
   IF #statErrorUserCleared = TRUE 
   THEN

       REGION Program

           //copy new value
           #statValues[0] := #statValues[1]; // -> n-2
           #statValues[1] := #statValues[2]; // -> n-1
           #statValues[2] := #statValues[3]; // -> n
           #statValues[3] := #statValues[4]; // -> n+1
           #statValues[4] := #value;         // -> n+2

           IF #statCount < 4
           THEN
               #status:= #STATUS_NOT_ENOUGH_VALUES;
               #statCount += 1;
               #statErrorAutoCleared := true;
           ELSE
               //calculate new smoothed value 
               //ẏ(n)=1/12deltaT*(y(n-2)-8y(n-1)+8y(n+1)-y(n+2))
               //1/12deltaT = 
               #statDerivatedValue := LREAL_TO_REAL(1.0 / (12.0*#deltaT)) * (#statValues[0] -8 * #statValues[1] + 8 * #statValues[3] - #statValues[4]);
               #statDone := true;
           END_IF;

       END_REGION
   END_IF;

   //----------------------------------------------------------------------------------------------
   //Write ouputs and error handling
   //----------------------------------------------------------------------------------------------
   //Error occured in request
   IF #statErrorAutoCleared
   THEN
       #statDone := FALSE;
       #statErrorUserCleared := FALSE;
       //Request finished
   ELSIF #statDone
   THEN
       #statErrorUserCleared := FALSE;
       #statErrorAutoCleared := FALSE;
       #status := #STATUS_EXECUTION_FINISHED;
       #derivatedValue := #statDerivatedValue;
       //Request in execution
   ELSE
       #status := #STATUS_SUBSEQUENT_CALL;
   END_IF;

   //Write static values to outputs
   #valid := #statDone;
   #busy := #statErrorUserCleared;
   #error := #statErrorAutoCleared;
   //----------------------------------------------------------------------------------------------

   //=============================================================================

   //----------------------------------------------------------------------------------------------
   //Check if FB is disabled
   IF NOT #enable
     AND #statEnableOld
   THEN

     //Error outputs are reset with falling edge of enable input
     #statErrorUserCleared := FALSE;
     #statErrorAutoCleared := FALSE;
     #error := FALSE;
     #status := #STATUS_NO_CALL;

     //Enable and busy are reset with falling edge of enable input
     #busy := FALSE;
     #busy := FALSE;

     //Set old value of enable for edge detection and end execution
     #statEnableOld := #enable;
     RETURN;

     //Check if FB is enabled
   ELSIF #enable
     AND NOT #statEnableOld
   THEN
     //reset static values
     #statCount := 0;
     #statValues[0] := 0.0;
     #statValues[1] := 0.0;
     #statValues[2] := 0.0;
     #statValues[3] := 0.0;
     #statValues[4] := 0.0;

     #derivatedValue := 0.0;
     #statNoValues := true;

     //Busy is set at rising edge of enable input
     #busy := TRUE;
     //Set status for first call
     #status := #STATUS_FIRST_CALL;
     //Set old value of enable for edge detection and end execution
     #statEnableOld := #enable;
     RETURN;

     //Check if user cleared error in FB occurred
   ELSIF #statErrorUserCleared


   THEN
     #busy := FALSE;
     //Set old value of enable for edge detection and end execution
     #statEnableOld := #enable;
     //No set of status necessary, because status already set when error occured
     RETURN;

     //Check if function block is disabled
   ELSIF NOT #enable
   THEN
     #busy := FALSE;
     #status := #STATUS_NO_CALL;
     //Set old value of enable for edge detection and end execution
     #statEnableOld := #enable;
     RETURN;

   ELSE
     //Detect edge for disabling
     #statEnableOld := #enable;
   END_IF;


   //----------------------------------------------------------------------------------------------
   //set Status "Not enough values" after reset
   IF #enable
     AND #statEnableOld
     AND #statNoValues
   THEN
     #status := #STATUS_NOT_ENOUGH_VALUES;
     #statErrorAutoCleared := true;
     #statNoValues := false;
   END_IF;

   // positive edge of insert detected 
   IF #insert
     AND NOT #statInsertOld
   THEN

     #statInsertOld := #insert;

     #statValues[0] := #statValues[1]; // -> n-2
     #statValues[1] := #statValues[2]; // -> n-1
     #statValues[2] := #statValues[3]; // -> n
     #statValues[3] := #statValues[4]; // -> n+1
     #statValues[4] := #value;         // -> n+2

     IF #statCount < 4 THEN
       #statCount += 1;
       #status := #STATUS_NOT_ENOUGH_VALUES;
       #statErrorAutoCleared := true;
     ELSE
       //calculate new smoothed value 
       //y(n)=1/35*(-3*y(n-2)+12*y(n-1)+17*y(n)+12*y(n+1)-3*y(n+2))
       //1/35 = 0.028571
       #derivatedValue := 0.028571 * (-3 * #statValues[0] + 12 * #statValues[1] + 17 * #statValues[2] + 12 * #statValues[3] - 3 * #statValues[4]);
     END_IF;
   ELSE

     #statInsertOld := #insert;
   END_IF;

   //----------------------------------------------------------------------------------------------
   //Error handling 
   //----------------------------------------------------------------------------------------------
   IF #statErrorUserCleared
   THEN
     #busy := FALSE;
     #busy := FALSE;
     #error := TRUE;

     RETURN;

   ELSIF #statErrorAutoCleared
   THEN
     #busy := FALSE;
     #busy := TRUE;
     #error := TRUE;

     RETURN;

   ELSE
     //Process normal output values
     #busy := TRUE;
     #error := FALSE;
     #status := #STATUS_SUBSEQUENT_CALL; //Set status for subsequent call
   END_IF;
   //----------------------------------------------------------------------------------------------
END_FUNCTION_BLOCK

FUNCTION "LGF_DifferenceQuotientFC" : Void   // FC3, SCL
{ S7_Optimized_Access := 'TRUE' }
VERSION : 0.1
   VAR_INPUT
      deltaT : Real;
   END_VAR
   VAR_OUTPUT
      error : Bool;
      status : Word;
   END_VAR
   VAR_IN_OUT
      values : Array[*] of Real;
      derivatedValues : Array[*] of Real;
   END_VAR
   VAR_TEMP
      tempLowerBound : DInt;
      tempUpperBound : DInt;
      tempNumberOfElements : DInt;
      tempLowerBoundOut : DInt;
      tempUpperBoundOut : DInt;
      tempNumberOfElementsOut : DInt;
      tempCount : Int;
      tempDivision : Real;
   END_VAR
   VAR CONSTANT
      STATUS_EXECUTION_FINISHED : Word := 16#0000;   // Execution finished without errors
      STATUS_NO_CALL : Word := 16#7000;   // No call of FB
      STATUS_NOT_ENOUGH_VALUES : Word := 16#9000;   // Not enough values. Min 5 Values are needed
      STATUS_ARRAYS_DIFFERENT : Word := 16#9001;   // Array values and Array derivatedValues need same size
   END_VAR
BEGIN
   //=============================================================================
   // SIEMENS AG
   // (c)Copyright 2017
   //-----------------------------------------------------------------------------
   // Library:       LGF (Library General Functions)
   // Tested with:   CPU1212C DC/DC/DC FW:V4.2
   // Engineering:   TIA Portal V15.1 
   // Restrictions:  -
   // Requirements:  PLC (S7-1200 / S7-1500)
   // Functionality: This function differentiates a signal 
   //-----------------------------------------------------------------------------
   // Change log table:
   // Version  Date        In charge / Changes applied
   // 01.00.00 23.11.2018  Siemens Industry Online Support
   //                      First released version
   //=============================================================================

   #error := false;

   REGION Program

       //check if size of arrays is ok
       #tempLowerBound := LOWER_BOUND(ARR := #values, DIM := 1);
       #tempUpperBound := UPPER_BOUND(ARR := #values, DIM := 1);

       #tempNumberOfElements := #tempUpperBound - #tempLowerBound;

       #tempLowerBoundOut := LOWER_BOUND(ARR := #derivatedValues, DIM := 1);
       #tempUpperBoundOut := UPPER_BOUND(ARR := #derivatedValues, DIM := 1);

       #tempNumberOfElementsOut := #tempUpperBoundOut - #tempLowerBoundOut;

       IF #tempNumberOfElementsOut <> #tempNumberOfElements
       THEN
         #error := true;
           #status := #STATUS_ARRAYS_DIFFERENT;
       ELSIF #tempNumberOfElements < 4
       THEN
           #status := #STATUS_NOT_ENOUGH_VALUES;
           #error := true;
       ELSE
           //ẏ(n)=1/12h*(y(n-2)-8y(n-1)+8y(n+1)-y(n+2))
           //h = deltaT

           #tempDivision := 1.0 / (12.0 * #deltaT);
           FOR #tempCount := #tempLowerBound + 2 TO #tempNumberOfElements-2 DO
             #derivatedValues[#tempCount] := #tempDivision * (#values[#tempCount-2] - 8 * #values[#tempCount -1] + 8 * #values[#tempCount + 1] - #values[#tempCount + 2]);
           END_FOR;

           //ẏ(n-2)=1/84h*(-125y(n-2)+136y(n-1)+48y(n)-88y(n+1)+29y(n+2))
           //h = deltaT
           #tempDivision := 1.0 / (84.0 * #deltaT);
           #derivatedValues[0] := #tempDivision * (-125 * #values[0] + 136 * #values[1] + 48 * #values[2] - 88 * #values[3] + 29* #values[4]);

           //ẏ(n-1)=1/84h*(-38y(n-2)-2y(n-1)+24y(n)+26y(n+1)-10y(n+2))
           //h = deltaT
           #derivatedValues[1] := #tempDivision * (-38 * #values[0] - 2 * #values[1] + 24 * #values[2] + 26 * #values[3] -10 * #values[4]);

           //ẏ(n+1)=1/84h(10y(n-2)-26y(n-1)-24y(n)+2y(n+1)+38y(n+2))
           //h = deltaT
           #derivatedValues[#tempUpperBound-1] := #tempDivision * (10 * #values[#tempUpperBound-4] - 26 * #values[#tempUpperBound-3]  -24 * #values[#tempUpperBound-2] +2 * #values[#tempUpperBound-1] + 38 * #values[#tempUpperBound]);

           //y(n-2)=1/84h(-29y(n-2)+88y(n-1)-48y(n)-136y(n+1)+125y(n+2))
           //h = deltaT
           #derivatedValues[#tempUpperBound] := #tempDivision * (-29 * #values[#tempUpperBound - 4] +88 * #values[#tempUpperBound - 3]  -48 * #values[#tempUpperBound - 2] -136 * #values[#tempUpperBound - 1] + 125 * #values[#tempUpperBound]);

           #status := #STATUS_EXECUTION_FINISHED;

       END_IF;
   END_REGION
END_FUNCTION

FUNCTION "LGF_AverageAndDeviation" : Void   // FC10006, SCL
{ S7_Optimized_Access := 'TRUE' }
   VAR_INPUT
      variableArray : Array[*] of LReal;   // Number series to be used for calculating
   END_VAR
   VAR_OUTPUT
      arithmeticAverage : LReal;   // Calculated Arithmetic average
      standardDeviation : LReal;   // Calculated Standard deviation
   END_VAR
   VAR_TEMP
      tempLowerBound : DInt;   // Temporary lower bound
      tempUpperBound : DInt;   // Temporary upper bound
      tempNumberOfElements : DInt;   // Temporary number of elements
      tempSizeCounter : Int;   // Temporary counter for loop
      tempArithmeticAverage : LReal;   // Temporary calculated Arithmetic average
      tempStandardDeviation : LReal;   // Temporary calculated Standard deviation
   END_VAR
   // Ret_Val : -
BEGIN
   //=============================================================================
   // SIEMENS AG
   // (c)Copyright 2017
   //-----------------------------------------------------------------------------
   // Library:       LGF (Library General Functions)
   // Tested with:   CPU1212C DC/DC/DC FW:V4.2
   // Engineering:   TIA Portal V14 Update 1
   // Restrictions:  -
   // Requirements:  PLC (S7-1200 / S7-1500)
   // Functionality: This function calculates the arithmetic average and the
   //                standard Deviation of a array of numbers
   //-----------------------------------------------------------------------------
   // Change log table:
   // Version  Date        In charge / Changes applied
   // 01.00.00 19.08.2015  Siemens Industry Online Support
   //                      First released version
   // 01.00.01 16.11.2015  Siemens Industry Online Support
   //                      Bug fix at WRONG_TYPE:  #error := true
   // 01.00.02 02.01.2017  Siemens Industry Online Support
   //                      Upgrade: TIA Portal V14 Update 1
   // 01.00.03 17.08.2018  Siemens Industry Online Support
   //                      Upgrade: TIA V15 Update 2
   // 01.00.04 23.11.2018  Siemens Industry Online Support
   //                      Upgrade: TIA V15.1
   // 02.00.00 25.01.2019  Siemens Industry Online Support
   //                      Data type changed from Variant to Array[*] of LReal
   //=============================================================================

   #tempLowerBound := LOWER_BOUND(ARR := #variableArray, DIM := 1);
   #tempUpperBound := UPPER_BOUND(ARR := #variableArray, DIM := 1);

   #tempNumberOfElements := #tempUpperBound - #tempLowerBound + 1;


   //------------------------------------------
   // Calculation of the arithmetic average
   //------------------------------------------
   #tempArithmeticAverage := 0;
   FOR #tempSizeCounter := #tempLowerBound TO #tempUpperBound DO
     #tempArithmeticAverage := #tempArithmeticAverage + #variableArray[#tempSizeCounter];
   END_FOR;

   #tempArithmeticAverage := #tempArithmeticAverage / DINT_TO_REAL(#tempNumberOfElements);

   //------------------------------------------
   //Calculation of the standardDeviation
   //------------------------------------------
   #tempStandardDeviation := 0;
   FOR #tempSizeCounter := #tempLowerBound TO #tempUpperBound DO
     #tempStandardDeviation := #tempStandardDeviation + SQR((#variableArray[#tempSizeCounter] - #tempArithmeticAverage));
   END_FOR;

   #tempStandardDeviation := #tempStandardDeviation / DINT_TO_REAL(#tempNumberOfElements);
   #tempStandardDeviation := SQRT(#tempStandardDeviation);

   #arithmeticAverage := #tempArithmeticAverage;
   #standardDeviation := #tempStandardDeviation;
END_FUNCTION

FUNCTION "LGF_SimpleSmoothingFC" : Void   // FC10012, SCL
{ S7_Optimized_Access := 'TRUE' }
VERSION : 0.1
   VAR_OUTPUT
      error : Bool;   // An error occurred during processing.
      status : Word;   // Outputs the status code of the processing (see table).
   END_VAR
   VAR_IN_OUT
      values : Array[*] of Real;   // Values that are to be included in the smoothing.
      smoothedValues : Array[*] of Real;   // The smoothed values.
   END_VAR
   VAR_TEMP
      tempCount : Int;   // Temporary count
      tempNumberOfElements : DInt;   // Temporary number of elements
      tempNumberOfElementsOut : DInt;   // Temporary number of elements out
      tempLowerBound : DInt;   // Temporary lower bound
      tempUpperBound : DInt;   // Temporary upper bound
      tempLowerBoundOut : DInt;   // Temporary lower bound out
      tempUpperBoundOut : DInt;   // Temporary upper bound out
   END_VAR
   VAR CONSTANT
      STATUS_EXECUTION_FINISHED : Word := 16#0000;   // Status: Execution finished without errors
      STATUS_NO_CALL : Word := 16#7000;   // Status: No call of FB
      STATUS_FIRST_CALL : Word := 16#7001;   // Status: First call of FB after enabling
      STATUS_SUBSEQUENT_CALL : Word := 16#7002;   // Status: Subsequent call of FB
      STATUS_NOT_ENOUGH_VALUES : Word := 16#9000;   // Status: Not enough values. Min 3 Values are needed
      STATUS_ARRAY_DIFFERENT : Word := 16#9001;   // Status: The Arraysizes are not equal
   END_VAR
BEGIN
   //=============================================================================
   // SIEMENS AG
   // (c)Copyright 2017
   //-----------------------------------------------------------------------------
   // Library:       LGF (Library General Functions)
   // Tested with:   CPU1212C DC/DC/DC FW:V4.2
   // Engineering:   TIA Portal V15.1 
   // Restrictions:  -
   // Requirements:  PLC (S7-1200 / S7-1500)
   // Functionality: This function calculates the smoothed values 
   //-----------------------------------------------------------------------------
   // Change log table:
   // Version  Date        In charge / Changes applied
   // 01.00.00 23.11.2018  Siemens Industry Online Support
   //                      First released version
   //=============================================================================

   #error := false;

   #tempLowerBound := LOWER_BOUND(ARR := #values, DIM := 1);
   #tempUpperBound := UPPER_BOUND(ARR := #values, DIM := 1);

   #tempNumberOfElements := #tempUpperBound - #tempLowerBound;

   #tempLowerBoundOut := LOWER_BOUND(ARR := #smoothedValues, DIM := 1);
   #tempUpperBoundOut := UPPER_BOUND(ARR := #smoothedValues, DIM := 1);

   #tempNumberOfElementsOut := #tempUpperBoundOut - #tempLowerBoundOut;

   IF #tempNumberOfElements <> #tempNumberOfElementsOut
   THEN
     #error := true;
     #status := #STATUS_ARRAY_DIFFERENT;
   ELSIF #tempNumberOfElements < 3
   THEN
     #status := #STATUS_NOT_ENOUGH_VALUES;
     #error := true;
   ELSE
     //y(Nsmoothed)= (y(n-1)+y(n)+y(n+1)) / 3
     FOR #tempCount := #tempLowerBound + 1 TO #tempUpperBound - 1 DO
       #smoothedValues[#tempCount] := (#values[#tempCount - 1] + #values[#tempCount] + #values[#tempCount + 1]) / 3;
     END_FOR;

   END_IF;
END_FUNCTION

FUNCTION "LGF_SmoothByPolynomFC" : Void   // FC10013, SCL
{ S7_Optimized_Access := 'TRUE' }
VERSION : 0.1
   VAR_OUTPUT
      error : Bool;   // An error occurred during processing.
      status : Word;   // Outputs the status code of the processing (see table).
   END_VAR
   VAR_IN_OUT
      values : Array[*] of Real;   // Values that are to be included in the smoothing.
      smoothedValues : Array[*] of Real;   // The smoothed values.
   END_VAR
   VAR_TEMP
      tempCount : Int;   // Temporary count
      tempNumberOfElements : DInt;   // Temporary number of elements
      tempNumberOfElementsOut : DInt;   // Temporary number of elements out
      tempLowerBound : DInt;   // Temporary lower bound
      tempUpperBound : DInt;   // Temporary upper bound
      tempLowerBoundOut : DInt;   // Temporary lower bound out
      tempUpperBoundOut : DInt;   // Temporary upper bound out
   END_VAR
   VAR CONSTANT
      STATUS_EXECUTION_FINISHED : Word := 16#0000;   // Status: Execution finished without errors
      STATUS_NO_CALL : Word := 16#7000;   // Status: No call of FB
      STATUS_NOT_ENOUGH_VALUES : Word := 16#9000;   // Status: Not enough values. Min 5 Values are needed
      STATUS_ARRAYS_DIFFERENT : Word := 16#9001;   // Status: The Arraysize of values and smoothedValues must be equal
   END_VAR
BEGIN
   //=============================================================================
   // SIEMENS AG
   // (c)Copyright 2017
   //-----------------------------------------------------------------------------
   // Library:       LGF (Library General Functions)
   // Tested with:   CPU1212C DC/DC/DC FW:V4.2
   // Engineering:   TIA Portal V15.1 
   // Restrictions:  -
   // Requirements:  PLC (S7-1200 / S7-1500)
   // Functionality: This function calculates the smoothed values by polynom
   //-----------------------------------------------------------------------------
   // Change log table:
   // Version  Date        In charge / Changes applied
   // 01.00.00 23.11.2018  Siemens Industry Online Support
   //                      First released version
   //=============================================================================

   #status := #STATUS_NO_CALL;
   #error := false;

   REGION Program
       #tempLowerBound := LOWER_BOUND(ARR := #values, DIM := 1);
       #tempUpperBound := UPPER_BOUND(ARR := #values, DIM := 1);

       #tempNumberOfElements := #tempUpperBound - #tempLowerBound;

       #tempLowerBoundOut := LOWER_BOUND(ARR := #smoothedValues, DIM := 1);
       #tempUpperBoundOut := UPPER_BOUND(ARR := #smoothedValues, DIM := 1);

       #tempNumberOfElementsOut := #tempUpperBoundOut - #tempLowerBoundOut;

       IF #tempNumberOfElements <> #tempNumberOfElementsOut
       THEN
         #status := #STATUS_ARRAYS_DIFFERENT;
           #error := true;
       ELSIF #tempNumberOfElements < 4
       THEN
           #status := #STATUS_NOT_ENOUGH_VALUES;
           #error := true;

       ELSE
           FOR #tempCount := #tempLowerBound + 2 TO #tempUpperBound - 2 DO

               //calculate new smoothed value 
               //y(n)=1/35*(-3*y(n-2)+12*y(n-1)+17*y(n)+12*y(n+1)-3*y(n+2))
               //1/35 = 0.028571
             #smoothedValues[#tempCount] := 0.028571 * (-3 * #values[#tempCount - 2] + 12 * #values[#tempCount - 1] + 17 * #values[#tempCount] + 12 * #values[#tempCount + 1] - 3 * #values[#tempCount + 2]);
           END_FOR;

           //calculate Replacementvalues for 0,1 and n-1,n

           //y(0) =1/70*(69*y(0)+4*y(1)-6*y(2)+4*y(3)-y(4))
           //1/70 = 0.014286
           #smoothedValues[#tempLowerBound] := 0.014286 * (69 * #values[#tempLowerBound] + 4 * #values[#tempLowerBound + 1] - 6 * #values[#tempLowerBound + 2] + 4 * #values[#tempLowerBound + 3] - #values[#tempLowerBound + 4]);

           //y(1) =2/70*(2*y(0)+27*y(1)+12*y(2)-8*y(3)+2*y(4))
           //2/70 = 0.028571
           #smoothedValues[#tempLowerBound + 1] := 0.028571 * (2 * #values[#tempLowerBound] + 27 * #values[#tempLowerBound + 1] + 12 * #values[#tempLowerBound + 2] - 8 * #values[#tempLowerBound + 3] + 2 * #values[#tempLowerBound + 4]);

           //y(n-1) =2/70*(2*y(n-4)-8*y(n-3)+12*y(n-2)+27*y(n-1)+2*y(n))
           //2/70 = 0.028571
           #smoothedValues[#tempUpperBound - 1] := 0.028571 * (2 * #values[#tempUpperBound - 4] - 8 * #values[#tempUpperBound - 3] + 12 * #values[#tempUpperBound - 2] + 27 * #values[#tempUpperBound - 1] + 2 * #values[#tempUpperBound]);

           //y(n) =1/70*(-y(n-4)+4*y(n-3)-6*y(n-2)+4*y(n-1)+69*y(n))
           //1/70 = 0.014286
           #smoothedValues[#tempUpperBound] := 0.014286 * (- #values[#tempUpperBound - 4] + 4 * #values[#tempUpperBound - 3] - 6 * #values[#tempUpperBound - 2] + 4 * #values[#tempUpperBound - 1] + 69 * #values[#tempUpperBound]);

           #status := #STATUS_EXECUTION_FINISHED;

       END_IF;
   END_REGION
END_FUNCTION

// folder: Phisical_functions/LGF/9 Measurement operations/LGF_RegressionLine

FUNCTION "LGF_RegressionLine" : Void   // FC8, SCL
{ S7_Optimized_Access := 'TRUE' }
VERSION : 0.1
   VAR_OUTPUT
      slope : LReal;   // Gradient of straight line
      intercept : LReal;   // The intersection with the Y axis
      error : Bool;   // An error occurred during processing
      status : Word;   // Outputs the status code of the processing
   END_VAR
   VAR_IN_OUT
      values : Array[*] of "LGF_typeRegressionLine";   // The data points are passed with their X- and Y-values
   END_VAR
   VAR_TEMP
      tempCount : DInt;   // Temporary count
      tempNumberOfElements : DInt;   // Temporary number of elements
      tempLowerBound : DInt;   // Temporary lower bound
      tempUpperBound : DInt;   // Temporary upper bound
      tempSumXY : LReal;   // Temporary sum XY
      tempSumX : LReal;   // Temporary sum X
      tempSumY : LReal;   // Temporary sum Y
      tempSumX2 : LReal;   // Temporary sum X2
      tempA : LReal;   // Temporary A
      tempB : LReal;   // Temporary B
      tempError : Bool;   // Temporary error
   END_VAR
   VAR CONSTANT
      STATUS_EXECUTION_FINISHED : Word := 16#0000;   // Execution finished without errors
      STATUS_NOT_ENOUGH_VALUES : Word := 16#9000;   // Not enough Values
   END_VAR
BEGIN
   //=============================================================================
   // SIEMENS AG
   // (c)Copyright 2017
   //-----------------------------------------------------------------------------
   // Library:       LGF (Library General Functions)
   // Tested with:   CPU1212C DC/DC/DC FW:V4.2
   // Engineering:   TIA Portal V15.1 
   // Restrictions:  -
   // Requirements:  PLC (S7-1200 / S7-1500)
   // Functionality: This function calculates the regression line 
   //-----------------------------------------------------------------------------
   // Change log table:
   // Version  Date        In charge / Changes applied
   // 01.00.00 23.11.2018  Siemens Industry Online Support
   //                      First released version
   //=============================================================================


   #error := false;

     //calculate number of elements
     #tempLowerBound := LOWER_BOUND(ARR := #values, DIM := 1);
     #tempUpperBound := UPPER_BOUND(ARR := #values, DIM := 1);

     #tempNumberOfElements := #tempUpperBound - #tempLowerBound + 1;

     //Not enough values 
     IF #tempNumberOfElements < 2
     THEN
       #tempError := true;
       #status := #STATUS_NOT_ENOUGH_VALUES;
       RETURN;
     END_IF;

     //caluclate sum of all needed values
     FOR #tempCount := #tempLowerBound TO #tempUpperBound
     DO
       //Sum of x(n) * y(n)
       #tempSumXY += #values[#tempCount].x * #values[#tempCount].y;
       //Sum of x(n) 
       #tempSumX += #values[#tempCount].x;
       //Sum of y(n)
       #tempSumY += #values[#tempCount].y;
       //Sum of x²(n)
       #tempSumX2 += SQR(#values[#tempCount].x);
     END_FOR;

     //b= (n* ∑(x(n)*y(n) - ( ∑x(n)* ∑y(n)))/
     //    (n* (∑x(n)^2) -(∑x(n)* ∑x(n)))
     #tempB := (#tempNumberOfElements * #tempSumXY - (#tempSumX * #tempSumY)) / (#tempNumberOfElements* #tempSumX2- (#tempSumX*#tempSumX));

     // a= Y-bX : X and Y are the average values of x and y
     #tempA := #tempSumY/ #tempNumberOfElements - (#tempB * (#tempSumX/ #tempNumberOfElements));


     // f(x)= a+b*x
     #slope := #tempB;
     #intercept := #tempA;

     #status := #STATUS_EXECUTION_FINISHED;
     #error := #tempError;
END_FUNCTION

// folder: Phisical_functions/LGF/99 Legacy

FUNCTION "LGF_CountFalInDWord" : Int   // FC10003, SCL
{ S7_Optimized_Access := 'TRUE' }
   VAR_INPUT
      dWordActCycle : DWord;
      dWordPrevCycle : DWord;
   END_VAR
   VAR_TEMP
      tempCount : Int;
   END_VAR
BEGIN
   //=============================================================================
   // SIEMENS AG
   // (c)Copyright 2017
   //-----------------------------------------------------------------------------
   // Library:       LGF (Library General Functions)
   // Tested with:   CPU1212C DC/DC/DC FW:V4.2
   // Engineering:   TIA Portal V14 Update 1
   // Restrictions:  -
   // Requirements:  PLC (S7-1200 / S7-1500)
   // Functionality: Detects and counts falling edges in variables of type DWORD
   //-----------------------------------------------------------------------------
   // Change log table:
   // Version  Date        In charge / Changes applied
   // 01.00.00 19.08.2015  Siemens Industry Online Support
   //                      First released version
   // 01.00.01 02.01.2017  Siemens Industry Online Support
   //                      Upgrade: TIA V14 Update 1
   // 01.00.02 17.08.2018  Siemens Industry Online Support
   //                      Upgrade: TIA V15 Update 2
   // 01.00.03 23.11.2018  Siemens Industry Online Support
   //                      Upgrade: TIA V15.1
   //=============================================================================

   // Initialization
   #tempCount := 0;

   //Byte 0
   //Bit                76543210765432107654321076543210         76543210765432107654321076543210
   IF ((#dWordActCycle AND DW#2#00000000000000000000000000000011) = DW#2#00000000000000000000000000000010) THEN
     #tempCount := #tempCount + 1;
   END_IF;
   //Bit                76543210765432107654321076543210         76543210765432107654321076543210
   IF ((#dWordActCycle AND DW#2#00000000000000000000000000000110) = DW#2#00000000000000000000000000000100) THEN
     #tempCount := #tempCount + 1;
   END_IF;
   //Bit                76543210765432107654321076543210         76543210765432107654321076543210
   IF ((#dWordActCycle AND DW#2#00000000000000000000000000001100) = DW#2#00000000000000000000000000001000) THEN
     #tempCount := #tempCount + 1;
   END_IF;
   //Bit                76543210765432107654321076543210         76543210765432107654321076543210
   IF ((#dWordActCycle AND DW#2#00000000000000000000000000011000) = DW#2#00000000000000000000000000010000) THEN
     #tempCount := #tempCount + 1;
   END_IF;
   //Bit                76543210765432107654321076543210         76543210765432107654321076543210
   IF ((#dWordActCycle AND DW#2#00000000000000000000000000110000) = DW#2#00000000000000000000000000100000) THEN
     #tempCount := #tempCount + 1;
   END_IF;
   //Bit             76543210765432107654321076543210         76543210765432107654321076543210
   IF ((#dWordActCycle AND DW#2#00000000000000000000000001100000) = DW#2#00000000000000000000000001000000) THEN
     #tempCount := #tempCount + 1;
   END_IF;
   //Bit             76543210765432107654321076543210         76543210765432107654321076543210
   IF ((#dWordActCycle AND DW#2#00000000000000000000000011000000) = DW#2#00000000000000000000000010000000) THEN
     #tempCount := #tempCount + 1;
   END_IF;
   //Bit                76543210765432107654321076543210         76543210765432107654321076543210
   IF ((#dWordActCycle AND DW#2#00000000000000000000000110000000) = DW#2#00000000000000000000000100000000) THEN
     #tempCount := #tempCount + 1;
   END_IF;

   //Byte 1
   //Bit                76543210765432107654321076543210         76543210765432107654321076543210
   IF ((#dWordActCycle AND DW#2#00000000000000000000001100000000) = DW#2#00000000000000000000001000000000) THEN
     #tempCount := #tempCount + 1;
   END_IF;
   //Bit                76543210765432107654321076543210         76543210765432107654321076543210
   IF ((#dWordActCycle AND DW#2#00000000000000000000011000000000) = DW#2#00000000000000000000010000000000) THEN
     #tempCount := #tempCount + 1;
   END_IF;
   //Bit                76543210765432107654321076543210         76543210765432107654321076543210
   IF ((#dWordActCycle AND DW#2#00000000000000000000110000000000) = DW#2#00000000000000000000100000000000) THEN
     #tempCount := #tempCount + 1;
   END_IF;
   //Bit                76543210765432107654321076543210         76543210765432107654321076543210
   IF ((#dWordActCycle AND DW#2#00000000000000000001100000000000) = DW#2#00000000000000000001000000000000) THEN
     #tempCount := #tempCount + 1;
   END_IF;
   //Bit                76543210765432107654321076543210         76543210765432107654321076543210
   IF ((#dWordActCycle AND DW#2#00000000000000000011000000000000) = DW#2#00000000000000000010000000000000) THEN
     #tempCount := #tempCount + 1;
   END_IF;
   //Bit                76543210765432107654321076543210         76543210765432107654321076543210
   IF ((#dWordActCycle AND DW#2#00000000000000000110000000000000) = DW#2#00000000000000000100000000000000) THEN
     #tempCount := #tempCount + 1;
   END_IF;
   //Bit                76543210765432107654321076543210         76543210765432107654321076543210
   IF ((#dWordActCycle AND DW#2#00000000000000001100000000000000) = DW#2#00000000000000001000000000000000) THEN
     #tempCount := #tempCount + 1;
   END_IF;
   //Bit             76543210765432107654321076543210         76543210765432107654321076543210
   IF ((#dWordActCycle AND DW#2#00000000000000011000000000000000) = DW#2#00000000000000010000000000000000) THEN
     #tempCount := #tempCount + 1;
   END_IF;

   //Byte 2
   //Bit                76543210765432107654321076543210         76543210765432107654321076543210
   IF ((#dWordActCycle AND DW#2#00000000000000110000000000000000) = DW#2#00000000000000100000000000000000) THEN
     #tempCount := #tempCount + 1;
   END_IF;
   //Bit                76543210765432107654321076543210         76543210765432107654321076543210
   IF ((#dWordActCycle AND DW#2#00000000000001100000000000000000) = DW#2#00000000000001000000000000000000) THEN
     #tempCount := #tempCount + 1;
   END_IF;
   //Bit                76543210765432107654321076543210         76543210765432107654321076543210
   IF ((#dWordActCycle AND DW#2#00000000000011000000000000000000) = DW#2#00000000000010000000000000000000) THEN
     #tempCount := #tempCount + 1;
   END_IF;
   //Bit             76543210765432107654321076543210         76543210765432107654321076543210
   IF ((#dWordActCycle AND DW#2#00000000000110000000000000000000) = DW#2#00000000000100000000000000000000) THEN
     #tempCount := #tempCount + 1;
   END_IF;
   //Bit                76543210765432107654321076543210         76543210765432107654321076543210
   IF ((#dWordActCycle AND DW#2#00000000001100000000000000000000) = DW#2#00000000001000000000000000000000) THEN
     #tempCount := #tempCount + 1;
   END_IF;
   //Bit                76543210765432107654321076543210         76543210765432107654321076543210
   IF ((#dWordActCycle AND DW#2#00000000011000000000000000000000) = DW#2#00000000010000000000000000000000) THEN
     #tempCount := #tempCount + 1;
   END_IF;
   //Bit                76543210765432107654321076543210         76543210765432107654321076543210
   IF ((#dWordActCycle AND DW#2#00000000110000000000000000000000) = DW#2#00000000100000000000000000000000) THEN
     #tempCount := #tempCount + 1;
   END_IF;
   //Bit                76543210765432107654321076543210         76543210765432107654321076543210
   IF ((#dWordActCycle AND DW#2#00000001100000000000000000000000) = DW#2#00000001000000000000000000000000) THEN
     #tempCount := #tempCount + 1;
   END_IF;

   //Byte 3
   //Bit                76543210765432107654321076543210         76543210765432107654321076543210
   IF ((#dWordActCycle AND DW#2#00000011000000000000000000000000) = DW#2#00000010000000000000000000000000) THEN
     #tempCount := #tempCount + 1;
   END_IF;
   //Bit                76543210765432107654321076543210         76543210765432107654321076543210
   IF ((#dWordActCycle AND DW#2#00000110000000000000000000000000) = DW#2#00000100000000000000000000000000) THEN
     #tempCount := #tempCount + 1;
   END_IF;
   //Bit                76543210765432107654321076543210         76543210765432107654321076543210
   IF ((#dWordActCycle AND DW#2#00001100000000000000000000000000) = DW#2#00001000000000000000000000000000) THEN
     #tempCount := #tempCount + 1;
   END_IF;
   //Bit                76543210765432107654321076543210         76543210765432107654321076543210
   IF ((#dWordActCycle AND DW#2#00011000000000000000000000000000) = DW#2#00010000000000000000000000000000) THEN
     #tempCount := #tempCount + 1;
   END_IF;
   //Bit                76543210765432107654321076543210         76543210765432107654321076543210
   IF ((#dWordActCycle AND DW#2#00110000000000000000000000000000) = DW#2#00100000000000000000000000000000) THEN
     #tempCount := #tempCount + 1;
   END_IF;
   //Bit                76543210765432107654321076543210         76543210765432107654321076543210
   IF ((#dWordActCycle AND DW#2#01100000000000000000000000000000) = DW#2#01000000000000000000000000000000) THEN
     #tempCount := #tempCount + 1;
   END_IF;
   //Bit                76543210765432107654321076543210         76543210765432107654321076543210
   IF ((#dWordActCycle AND DW#2#11000000000000000000000000000000) = DW#2#10000000000000000000000000000000) THEN
     #tempCount := #tempCount + 1;
   END_IF;
   //Bit                 76543210765432107654321076543210         76543210765432107654321076543210
   IF (((#dWordActCycle AND DW#2#10000000000000000000000000000000) = DW#2#00000000000000000000000000000000)
     AND ((#dWordPrevCycle AND DW#2#00000000000000000000000000000001) = DW#2#00000000000000000000000000000001))
   THEN
     #tempCount := #tempCount + 1;
   END_IF;

   //Output
   #LGF_CountFalInDWord := #tempCount;
END_FUNCTION

FUNCTION "LGF_CountRisInDWord" : Int   // FC10004, SCL
{ S7_Optimized_Access := 'TRUE' }
   VAR_INPUT
      dWordActCycle : DWord;
      dWordPrevCycle : DWord;
   END_VAR
   VAR_TEMP
      tempCount : Int;
   END_VAR
BEGIN
   //=============================================================================
   // SIEMENS AG
   // (c)Copyright 2017
   //-----------------------------------------------------------------------------
   // Library:       LGF (Library General Functions)
   // Tested with:   CPU1212C DC/DC/DC FW:V4.2
   // Engineering:   TIA Portal V14 Update 1
   // Restrictions:  -
   // Requirements:  PLC (S7-1200 / S7-1500)
   // Functionality: Detects rising edges in variables of type DWORD
   //-----------------------------------------------------------------------------
   // Change log table:
   // Version  Date        In charge / Changes applied
   // 01.00.00 19.08.2015  Siemens Industry Online Support
   //                      First released version
   // 01.00.01 02.01.2017  Siemens Industry Online Support
   //                      Upgrade: TIA V14 Update 1
   // 01.00.02 17.08.2018  Siemens Industry Online Support
   //                      Upgrade: TIA V15 Update 2
   // 01.00.03 23.11.2018  Siemens Industry Online Support
   //                      Upgrade: TIA V15.1
   //=============================================================================

   // Initialization
   #tempCount := 0;

   //Byte 0
   //Bit                76543210765432107654321076543210         76543210765432107654321076543210
   IF ((#dWordActCycle AND DW#2#00000000000000000000000000000011) = DW#2#00000000000000000000000000000001) THEN
     #tempCount := #tempCount + 1;
   END_IF;
   //Bit                76543210765432107654321076543210         76543210765432107654321076543210
   IF ((#dWordActCycle AND DW#2#00000000000000000000000000000110) = DW#2#00000000000000000000000000000010) THEN
     #tempCount := #tempCount + 1;
   END_IF;
   //Bit                76543210765432107654321076543210         76543210765432107654321076543210
   IF ((#dWordActCycle AND DW#2#00000000000000000000000000001100) = DW#2#00000000000000000000000000000100) THEN
     #tempCount := #tempCount + 1;
   END_IF;
   //Bit                76543210765432107654321076543210         76543210765432107654321076543210
   IF ((#dWordActCycle AND DW#2#00000000000000000000000000011000) = DW#2#00000000000000000000000000001000) THEN
     #tempCount := #tempCount + 1;
   END_IF;
   //Bit                76543210765432107654321076543210         76543210765432107654321076543210
   IF ((#dWordActCycle AND DW#2#00000000000000000000000000110000) = DW#2#00000000000000000000000000010000) THEN
     #tempCount := #tempCount + 1;
   END_IF;
   //Bit                76543210765432107654321076543210         76543210765432107654321076543210
   IF ((#dWordActCycle AND DW#2#00000000000000000000000001100000) = DW#2#00000000000000000000000000100000) THEN
     #tempCount := #tempCount + 1;
   END_IF;
   //Bit                76543210765432107654321076543210         76543210765432107654321076543210
   IF ((#dWordActCycle AND DW#2#00000000000000000000000011000000) = DW#2#00000000000000000000000001000000) THEN
     #tempCount := #tempCount + 1;
   END_IF;
   //Bit                76543210765432107654321076543210         76543210765432107654321076543210
   IF ((#dWordActCycle AND DW#2#00000000000000000000000110000000) = DW#2#00000000000000000000000010000000) THEN
     #tempCount := #tempCount + 1;
   END_IF;

   //Byte 1
   //Bit                76543210765432107654321076543210         76543210765432107654321076543210
   IF ((#dWordActCycle AND DW#2#00000000000000000000001100000000) = DW#2#00000000000000000000000100000000) THEN
     #tempCount := #tempCount + 1;
   END_IF;
   //Bit                76543210765432107654321076543210         76543210765432107654321076543210
   IF ((#dWordActCycle AND DW#2#00000000000000000000011000000000) = DW#2#00000000000000000000001000000000) THEN
     #tempCount := #tempCount + 1;
   END_IF;
   //Bit                76543210765432107654321076543210         76543210765432107654321076543210
   IF ((#dWordActCycle AND DW#2#00000000000000000000110000000000) = DW#2#00000000000000000000010000000000) THEN
     #tempCount := #tempCount + 1;
   END_IF;
   //Bit                76543210765432107654321076543210         76543210765432107654321076543210
   IF ((#dWordActCycle AND DW#2#00000000000000000001100000000000) = DW#2#00000000000000000000100000000000) THEN
     #tempCount := #tempCount + 1;
   END_IF;
   //Bit                76543210765432107654321076543210         76543210765432107654321076543210
   IF ((#dWordActCycle AND DW#2#00000000000000000011000000000000) = DW#2#00000000000000000001000000000000) THEN
     #tempCount := #tempCount + 1;
   END_IF;
   //Bit                76543210765432107654321076543210         76543210765432107654321076543210
   IF ((#dWordActCycle AND DW#2#00000000000000000110000000000000) = DW#2#00000000000000000010000000000000) THEN
     #tempCount := #tempCount + 1;
   END_IF;
   //Bit                76543210765432107654321076543210         76543210765432107654321076543210
   IF ((#dWordActCycle AND DW#2#00000000000000001100000000000000) = DW#2#00000000000000000100000000000000) THEN
     #tempCount := #tempCount + 1;
   END_IF;
   //Bit                76543210765432107654321076543210         76543210765432107654321076543210
   IF ((#dWordActCycle AND DW#2#00000000000000011000000000000000) = DW#2#00000000000000001000000000000000) THEN
     #tempCount := #tempCount + 1;
   END_IF;

   //Byte 2
   //Bit                76543210765432107654321076543210         76543210765432107654321076543210
   IF ((#dWordActCycle AND DW#2#00000000000000110000000000000000) = DW#2#00000000000000010000000000000000) THEN
     #tempCount := #tempCount + 1;
   END_IF;
   //Bit                76543210765432107654321076543210         76543210765432107654321076543210
   IF ((#dWordActCycle AND DW#2#00000000000001100000000000000000) = DW#2#00000000000000100000000000000000) THEN
     #tempCount := #tempCount + 1;
   END_IF;
   //Bit                76543210765432107654321076543210         76543210765432107654321076543210
   IF ((#dWordActCycle AND DW#2#00000000000011000000000000000000) = DW#2#00000000000001000000000000000000) THEN
     #tempCount := #tempCount + 1;
   END_IF;
   //Bit                76543210765432107654321076543210         76543210765432107654321076543210
   IF ((#dWordActCycle AND DW#2#00000000000110000000000000000000) = DW#2#00000000000010000000000000000000) THEN
     #tempCount := #tempCount + 1;
   END_IF;
   //Bit                76543210765432107654321076543210         76543210765432107654321076543210
   IF ((#dWordActCycle AND DW#2#00000000001100000000000000000000) = DW#2#00000000000100000000000000000000) THEN
     #tempCount := #tempCount + 1;
   END_IF;
   //Bit                76543210765432107654321076543210         76543210765432107654321076543210
   IF ((#dWordActCycle AND DW#2#00000000011000000000000000000000) = DW#2#00000000001000000000000000000000) THEN
     #tempCount := #tempCount + 1;
   END_IF;
   //Bit                76543210765432107654321076543210         76543210765432107654321076543210
   IF ((#dWordActCycle AND DW#2#00000000110000000000000000000000) = DW#2#00000000010000000000000000000000) THEN
     #tempCount := #tempCount + 1;
   END_IF;
   //Bit                76543210765432107654321076543210         76543210765432107654321076543210
   IF ((#dWordActCycle AND DW#2#00000001100000000000000000000000) = DW#2#00000000100000000000000000000000) THEN
     #tempCount := #tempCount + 1;
   END_IF;

   //Byte 3
   //Bit                76543210765432107654321076543210         76543210765432107654321076543210
   IF ((#dWordActCycle AND DW#2#00000011000000000000000000000000) = DW#2#00000001000000000000000000000000) THEN
     #tempCount := #tempCount + 1;
   END_IF;
   //Bit                76543210765432107654321076543210         76543210765432107654321076543210
   IF ((#dWordActCycle AND DW#2#00000110000000000000000000000000) = DW#2#00000010000000000000000000000000) THEN
     #tempCount := #tempCount + 1;
   END_IF;
   //Bit                76543210765432107654321076543210         76543210765432107654321076543210
   IF ((#dWordActCycle AND DW#2#00001100000000000000000000000000) = DW#2#00000100000000000000000000000000) THEN
     #tempCount := #tempCount + 1;
   END_IF;
   //Bit                76543210765432107654321076543210         76543210765432107654321076543210
   IF ((#dWordActCycle AND DW#2#00011000000000000000000000000000) = DW#2#00001000000000000000000000000000) THEN
     #tempCount := #tempCount + 1;
   END_IF;
   //Bit                76543210765432107654321076543210         76543210765432107654321076543210
   IF ((#dWordActCycle AND DW#2#00110000000000000000000000000000) = DW#2#00010000000000000000000000000000) THEN
     #tempCount := #tempCount + 1;
   END_IF;
   //Bit                76543210765432107654321076543210         76543210765432107654321076543210
   IF ((#dWordActCycle AND DW#2#01100000000000000000000000000000) = DW#2#00100000000000000000000000000000) THEN
     #tempCount := #tempCount + 1;
   END_IF;
   //Bit                76543210765432107654321076543210         76543210765432107654321076543210
   IF ((#dWordActCycle AND DW#2#11000000000000000000000000000000) = DW#2#01000000000000000000000000000000) THEN
     #tempCount := #tempCount + 1;
   END_IF;
   //Bit                 76543210765432107654321076543210         76543210765432107654321076543210
   IF (((#dWordActCycle AND DW#2#10000000000000000000000000000000) = DW#2#10000000000000000000000000000000)
     AND ((#dWordPrevCycle AND DW#2#00000000000000000000000000000001) = DW#2#00000000000000000000000000000000))
   THEN
     #tempCount := #tempCount + 1;
   END_IF;

   //Output
   #LGF_CountRisInDWord := #tempCount;
END_FUNCTION

(* ===== HMI "HMI_RT_1" =====
system functions are stored by id; their names below are inferred from use
connection "HMI_Connection_1": ETHERNET, S7_1200_OMS

